
                                   REGION "GET FROM HMI"
                                       #dzLabel := #settings.viewingStation.dzData.value;
                                   END_REGION

                                   REGION "WRITE TO STATION PARAMETER"
                                       #stations.me[#i].dropZone := WSTRING_TO_USINT(#dzLabel);
                                   END_REGION

                               END_IF;
                           END_REGION

                           REGION "ON LINE LABEL INPUT"
                               IF #lineEntered THEN

                                   REGION "GET FROM HMI"
                                       #lineLabel := #settings.viewingStation.lineData.value;
                                   END_REGION

                                   REGION "WRITE TO STATION PARAMETER"
                                       #stations.me[#i].line := #lineLabel;
                                   END_REGION

                               END_IF;
                           END_REGION

                       END_IF;
                   END_REGION

               END_FOR;
           END_REGION

       END_IF;
   END_REGION
END_FUNCTION

FUNCTION "Animate Button Details" : Void   // FC19, SCL
{ S7_Optimized_Access := 'TRUE' }
VERSION : 0.1
   VAR_INPUT
      stations : "Stations";
   END_VAR
   VAR_IN_OUT
      settings : "Settings";
   END_VAR
   VAR_TEMP
      animate : USInt;
      btnCount : Int;
      btnSelected : Bool;
      deselected : USInt;
      i : Int;
      invisible : USInt;
      pBtn : Int;
      selected : USInt;
      selStnCount : Int;
      selStnNumber : Int;
   END_VAR
BEGIN
   REGION "COPY TO LOCAL"
       #btnCount := "ptsPerStn";
       #deselected := "BgGray";
       #invisible := "invisible";
       #selected := "BgLTe";
       #selStnCount := #settings.#stations.selCount;
       #selStnNumber := #settings.stations.selNumber;
   END_REGION

   REGION "ENABLE"
       IF #selStnCount >= 1 THEN

           REGION "SHOW BUTTON DETAILS"
               #animate := #deselected;
           END_REGION

       END_IF;
   END_REGION

   REGION "DISABLE"
       IF #selStnCount = 0 THEN

           REGION "HIDE BUTTON DETAILS"
               #animate := #invisible;
           END_REGION

       END_IF;
   END_REGION

   REGION "APPLY ANIMATION"
       FOR #i := 0 TO #btnCount DO

           REGION "CALCULATE BUTTON POINTER"
               #pBtn := "Pointer Calc: Button Details"(#i);
           END_REGION

           REGION "WHILE Station SELECTED"
               IF #selStnCount <> 0 THEN

                   REGION "COPY TO LOCAL"
                       #btnSelected := #stations.me[#selStnNumber].settings.btnSelection[#pBtn];
                   END_REGION

                   REGION "ANIMATE BUTTON SELECTION

                       REGION "SELECTED"
                           IF #btnSelected THEN
                               #animate := #selected;
                           END_IF;
                       END_REGION

                       REGION "NOT SELECTED"
                           IF NOT #btnSelected THEN
                               #animate := #deselected;
                           END_IF;
                       END_REGION

                   END_REGION

               END_IF;
           END_REGION


           REGION "SEND TO HMI"
               #settings.viewingStation.btns[#i].label.animate := #animate;
               #settings.viewingStation.btns[#i].alloted.animate := #animate;
               #settings.viewingStation.btns[#i].critical.animate := #animate;
               #settings.viewingStation.btns[#i].partNumber.animate := #animate;
           END_REGION

       END_FOR;
   END_REGION
END_FUNCTION

FUNCTION "Populate Station Name" : WString   // FC20, SCL
{ S7_Optimized_Access := 'TRUE' }
VERSION : 0.1
   VAR_INPUT
      line : WString;
      dropZone : USInt;
   END_VAR
BEGIN
   #"Populate Station Name" := CONCAT_WSTRING(IN1 := #line,
                                              IN2 := wstring#' ',
                                              IN3 := "Strip Sign"(USINT_TO_WSTRING(#dropZone)));
END_FUNCTION

FUNCTION "Pointer Calc: Button Details" : Int   // FC21, SCL
{ S7_Optimized_Access := 'TRUE' }
VERSION : 0.1
   VAR_INPUT
      index : Int;
   END_VAR
   VAR_TEMP
      val : Int;
   END_VAR
BEGIN
   IF #index MOD 2 = 0 THEN
       #val := 7 - #index / 2;
   END_IF;

   IF #index MOD 2 <> 0 THEN
       #val := 3 - #index / 2;
   END_IF;

   #"Pointer Calc: Button Details" := #val;
END_FUNCTION

FUNCTION "Buffer Part Req Log Row: Generate" : "Part Req Log Row"   // FC22, SCL
{ S7_Optimized_Access := 'TRUE' }
VERSION : 0.1
   VAR_INPUT
      address : Int;
      "type" : Int;
   END_VAR
   VAR_TEMP
      retVal : Int;
   END_VAR
BEGIN
   REGION "ADDRESS"
       #"Buffer Part Req Log Row: Generate".address := #address;
   END_REGION

   REGION "REQUEST TYPE"
       #"Buffer Part Req Log Row: Generate".reqType := #type;
   END_REGION

   REGION "TIME STAMP"
       #retVal := RD_SYS_T(#"Buffer Part Req Log Row: Generate".timeStamp);
   END_REGION
END_FUNCTION

FUNCTION "Sim to Global" : Void   // FC23, SCL
{ S7_Optimized_Access := 'TRUE' }
VERSION : 0.1
   VAR_INPUT
      simStations : "Simulated Stations";
   END_VAR
   VAR_IN_OUT
      stations : "Stations";
   END_VAR
   VAR_TEMP
      btnCount : Int;
      firstStn : Int;
      i : Int;
      j : Int;
      pSim : Int;
      pStn : Int;
      simKP8Count : Int;
      stnCount : Int;
   END_VAR
BEGIN
   REGION "COPY TO LOCAL"
       #btnCount := "ptsPerStn";
       #firstStn := #simStations.firstStn;
       #simKP8Count := "simKP8Count";
       #stnCount := "stnCount";
   END_REGION

   REGION "FOR EACH STATION"
       FOR #i := 0 TO #simKP8Count DO

           REGION "CALCULATE POINTER"
               #pStn := #i + #firstStn;
               #pSim := #i;
           END_REGION

           REGION "UPPER LIMIT ROLL OVER"
               IF #pStn > #stnCount THEN
                   #pStn := #firstStn + #i - #stnCount - 1;
               END_IF;
           END_REGION

           REGION "COPY SIMULATED PRESSES"
               #stations.me[#pStn].kp8In := #simStations.me[#pSim].btn.actuate;
           END_REGION

       END_FOR;
   END_REGION
END_FUNCTION

FUNCTION "Pointer Calc: KP8 Labels" : Int   // FC25, SCL
{ S7_Optimized_Access := 'TRUE' }
VERSION : 0.1
   VAR_INPUT
      index : Int;
   END_VAR
   VAR_TEMP
      val : Int;
   END_VAR
BEGIN
   IF #index >= 4 THEN
       #val := 7 - (#index - 4) * 2;
   END_IF;

   IF #index <= 3 THEN
       #val := 8 - #index * 2;
   END_IF;

   #"Pointer Calc: KP8 Labels" := #val;
END_FUNCTION

FUNCTION "KP8 Color to Sim Animation" : USInt   // FC26, SCL
{ S7_Optimized_Access := 'TRUE' }
VERSION : 0.1
   VAR_INPUT
      kp8Color : DWord;
      btnNumber : Int;
   END_VAR
   VAR_TEMP
      animate : USInt;
      blue : USInt;
      colorDWord : DWord;
      colorInt : DInt;
      green : USInt;
      off : USInt;
      red : USInt;
      white : USInt;
      yellow : USInt;
   END_VAR
   VAR CONSTANT
      blueMask : DInt := 16#0000_0100;
      btnMask : DInt := 16#0101_0100;
      greenMask : DInt := 16#0001_0000;
      offMask : DInt := 16#0000_0000;
      redMask : DInt := 16#0100_0000;
      whiteMask : DInt := 16#0101_0100;
      yellowMask : DInt := 16#0101_0000;
   END_VAR
BEGIN
   REGION "COPY TO LOCAL"
       #blue := "BgLBl";
       #green := "BgLGr";
       #off := "BgGray";
       #red := "BgLRd";
       #white := "BgWh";
       #yellow := "BgLYe";
   END_REGION

   REGION "ISOLATE BUTTON COLOR"
       #colorDWord := SHR_DWORD(IN := #kp8Color,N := INT_TO_ULINT(#btnNumber));
       #colorDWord := #colorDWord AND #btnMask;
       #colorInt := DWORD_TO_DINT(#colorDWord);
   END_REGION

   REGION "DETERMINE ANIMATION"
       CASE #colorInt OF
           #blueMask:
               #animate := #blue;
           #greenMask:
               #animate := #green;
           #redMask:
               #animate := #red;
           #whiteMask:
               #animate := #white;
           #yellowMask:
               #animate := #yellow;
           ELSE
               #animate := #off;
       END_CASE;
   END_REGION

   REGION "RETURN VALUE"
       #"KP8 Color to Sim Animation" := #animate;
   END_REGION
END_FUNCTION

FUNCTION "Recipe Nav Button" : Void   // FC32, SCL
{ S7_Optimized_Access := 'TRUE' }
VERSION : 0.1
   VAR_INPUT
      visRows : Int;
      actuate : Bool;
      maxRows : Int;
      btnNum : Int;
   END_VAR
   VAR_IN_OUT
      recipeSelectScreen : "HSS: Menu Selection Screen";
   END_VAR
   VAR_TEMP
      eval : "HSS: Menu Selection Screen";
      color : Int;
   END_VAR
BEGIN
   REGION "COPY TO LOCAL"
       #eval := #recipeSelectScreen;
   END_REGION


   REGION "NARROW"
       IF #maxRows > #visRows THEN
           #color := "BgGray";
       END_IF;
   END_REGION


   REGION "WIDE"
       IF #maxRows <= #visRows THEN
           #color := "invisible";
       END_IF;
   END_REGION


   REGION "ROW COUNT INDEPENDENT"
       IF #actuate THEN
           #color := "BgLTe";
       END_IF;
   END_REGION


   REGION "DRAW"
       #eval.animate[#btnNum] := #color;
   END_REGION


   REGION "COPY TO GLOBAL"
       #recipeSelectScreen := #eval;
   END_REGION
END_FUNCTION

FUNCTION "LRUD KP8 Remap" : Int   // FC35, SCL
{ S7_Optimized_Access := 'TRUE' }
VERSION : 0.1
   VAR_INPUT
      btnNum : Int;
      mode : Int;   // 1 = KP8; 2 = KTP700
   END_VAR
   VAR_TEMP
      output : Int;
   END_VAR
   VAR CONSTANT
      kp8 : Int := 1;
      ktp700 : Int := 2;
   END_VAR
BEGIN
   IF #btnNum >= 4 THEN
       #output := (7 - #btnNum) * 2;
   END_IF;

   IF #btnNum <= 3 THEN
       #output := (3 - #btnNum) * 2 + 1;
   END_IF;

   #"LRUD KP8 Remap" := #output;
END_FUNCTION

// folder: Unsorted/Main HMI/Network Diagnostics

FUNCTION_BLOCK "NetDiag: Get IPs"   // FB27, SCL
{ S7_Optimized_Access := 'TRUE' }
VERSION : 0.1
   VAR_OUTPUT
      error : Bool := FALSE;   // Rising edge informs that an error occurred during the execution of the FB
      status : Word := 16#0000;   // Current status of FB
      statusID : Word := 16#0;   // Current status ID of calling instruction
   END_VAR
   VAR_IN_OUT
      ioSystemData : "UserDiag_typeIOSystem";   // IO-System diagnostics data
   END_VAR
   VAR
      statError : Bool := FALSE;   // Static value for output error
      statStatus : Word := 16#0000;   // Static value for output status
      statStatusID : Word := 16#0;   // Static value for output statusID
      instGetStationInfo : GetStationInfo;   // Instance of GetStationInfo
      statFirstDeviceFlag : Bool := TRUE;   // Help tag for the first device in the linked list
      statDeviceIndex : Int := 0;   // Device/slave index
   END_VAR
   VAR_TEMP
      tempIP : IF_CONF_v4;   // Temporary IP address
   END_VAR
   VAR CONSTANT
      STATUS_EXECUTION_FINISHED : Word := 16#0000;   // Execution finished without errors
      ID_GET_STATION_INFO : Word := 12;   // StatusID during GetStationInfo command
      MODE_IPV4 : UInt := 1;   // Address parameter according to IPv4
      LAST_DEVICE : Int := -1;   // No next device
   END_VAR
BEGIN
   //=============================================================================
   //SIEMENS AG
   //(c)Copyright 2015 All Rights Reserved
   //-----------------------------------------------------------------------------
   //Library: 
   //Tested with: S7-1516-3 PN/DP FW 2.5
   //Engineering: TIA Portal V15
   //Restrictions: Call in cyclic OB
   //Requirements: -
   //Functionality: Get IP address of IO devices
   //-----------------------------------------------------------------------------
   //Change log table:
   //Version  Date       Expert in charge                Changes applied
   //01.00.00 20.12.2017 Siemens Industry Online Support First released version
   //=============================================================================

   //=============================================================================
   // Go through existing devices and get IP address
   //=============================================================================
   // Initialize the pointer for the first run 
   IF (#statFirstDeviceFlag = TRUE)
   THEN
       #statDeviceIndex := #ioSystemData.firstDevice;
       #statFirstDeviceFlag := FALSE;
   END_IF;

   // Check and store the IP address, if the device is existing
   // GetStationInfo is an acyclic instruction. In the FB, the
   // instruction has to be repeated until it is done or error
   IF ((#ioSystemData.number >= 100)
       AND (#ioSystemData.number <= 115)
       AND (#ioSystemData.devices[#statDeviceIndex].exists = TRUE)
       AND (#ioSystemData.devices[#statDeviceIndex].ipAddress.ADDR[1] = 0))
   THEN
       // Get IP address of each decive in PN System
       #instGetStationInfo(REQ := TRUE,
                           LADDR := #ioSystemData.devices[#statDeviceIndex].hardwareId,
                           MODE := #MODE_IPV4,
                           DATA := #tempIP);

       IF (#instGetStationInfo.ERROR = TRUE)
       THEN
           // Error handling
           #statStatus := #instGetStationInfo.STATUS;
           #statStatusID := #ID_GET_STATION_INFO;
           #statError := TRUE;

           // Everything is ok --> Copy IP address    
       ELSIF (#instGetStationInfo.DONE = TRUE)
       THEN
           #ioSystemData.devices[#statDeviceIndex].ipAddress := #tempIP.InterfaceAddress;

           // Initialize the pointer for the next run
           #statDeviceIndex := #ioSystemData.devices[#statDeviceIndex].nextDevice;
       ELSE
           ;
       END_IF;
   ELSE
       // Initialize the pointer for the next run
       #statDeviceIndex := #ioSystemData.devices[#statDeviceIndex].nextDevice;
   END_IF;

   // Check last device
   IF (#statDeviceIndex = #LAST_DEVICE)
   THEN
       #statDeviceIndex := #ioSystemData.firstDevice;
   END_IF;

   // Write static values to outputs
   #error := #statError;
   #status := #statStatus;
   #statusID := #statStatusID;
END_FUNCTION_BLOCK

FUNCTION_BLOCK "NetDiag: Coordinate"   // FB28, LAD
{ S7_Optimized_Access := 'TRUE' }
VERSION : 0.1
// //============================================================================
// //SIEMENS AG
// //(c)Copyright 2017 All Rights Reserved
// //-----------------------------------------------------------------------------
// //Library: -
// //Tested with: S7-1516-3 PN/DP FW 2.5
// //Engineering: TIA Portal V15
// //Restrictions: -
// //Requirements: -
// //Functionality: Main FB for diagnostics
// //-----------------------------------------------------------------------------
// //Change log table:
// //Version  Date              Expert in charge                               Changes applied
// //01.00.00 25.04.2017 Siemens Industry Online Support First released version
// //01.01.00 01.12.2017 Siemens Industry Online Support Renamed in "UserDiag_Diagnostics"
// //                                                                                                    Check Flag "startDiag"
// //============================================================================
   VAR_IN_OUT
      startDiag : Bool := false;   // Startflag for diagnostic
      plcData : "UserDiag_typePLC";   // PLC diagnostics data
      ioSystemData : Array[1.."USERDIAG_IO_SYSTEMS_UPPER_LIM"] of "UserDiag_typeIOSystem";   // IO-System diagnostics data
   END_VAR
   VAR
      instPLCChk : "NetDiag: Check PLC";   // Instance of "UserDiag_PLCCheck"
      instIOSysChk : "NetDiag: IO Systems";   // Instance of "UserDiag_IOSystemCheck"
   END_VAR
BEGIN

REGION Network 1: Check Startflag for diagnostic
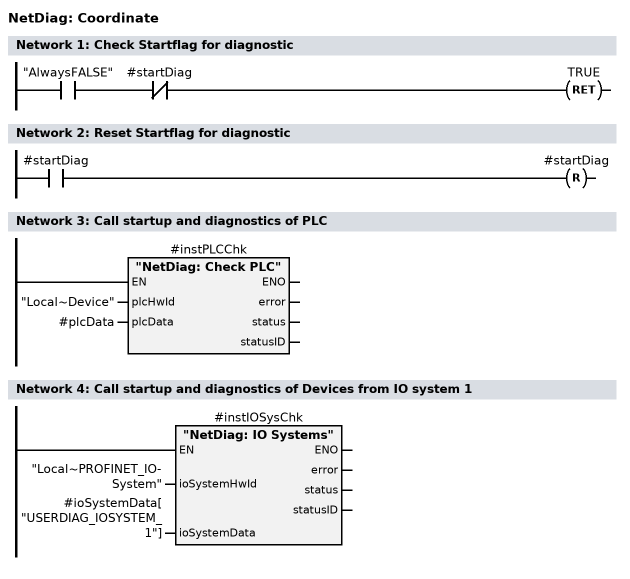
   IF "AlwaysFALSE" AND NOT #startDiag THEN
       ENO := TRUE;
       RETURN;
   END_IF;
END_REGION

REGION Network 2: Reset Startflag for diagnostic
   RUNG wire#powerrail
      Contact( #startDiag )
      R_Coil( #startDiag )
   END_RUNG
   // the same network as SCL:
   IF #startDiag THEN #startDiag := FALSE; END_IF;
END_REGION

REGION Network 3: Call startup and diagnostics of PLC
   RUNG wire#powerrail
      #instPLCChk(plcHwId := "Local~Device", plcData := #plcData, error =>, status =>, statusID =>)
   END_RUNG
   // the same network as SCL:
   #instPLCChk(plcHwId := "Local~Device", plcData := #plcData);   // "NetDiag: Check PLC"
END_REGION

REGION Network 4: Call startup and diagnostics of Devices from IO system 1
   RUNG wire#powerrail
      #instIOSysChk(ioSystemHwId := "Local~PROFINET_IO-System", ioSystemData := #ioSystemData["USERDIAG_IOSYSTEM_1"], error =>, status =>, statusID =>)
   END_RUNG
   // the same network as SCL:
   #instIOSysChk(ioSystemHwId := "Local~PROFINET_IO-System",   // "NetDiag: IO Systems"
                 ioSystemData := #ioSystemData["USERDIAG_IOSYSTEM_1"]);
END_REGION
END_FUNCTION_BLOCK

FUNCTION_BLOCK "NetDiag: Check PLC"   // FB29, SCL
{ S7_Optimized_Access := 'TRUE' }
VERSION : 0.1
   VAR_INPUT
      plcHwId : Hw_Device := 0;   // Hardware ID
   END_VAR
   VAR_OUTPUT
      error : Bool := FALSE;   // Rising edge informs that an error occurred during the execution of the FB
      status : Word := 16#0000;   // Current status of FB
      statusID : Word := 16#0;   // Current status ID of calling instruction
   END_VAR
   VAR_IN_OUT
      plcData : "UserDiag_typePLC";   // PLC diagnostics data
   END_VAR
   VAR
      statError : Bool := FALSE;   // Static value for output error
      statStatus : Word := 16#0000;   // Static value for output status
      statStatusID : Word := 16#0;   // Static value for output statusID
      statGeoAddr : GEOADDR;   // Slot information
      statGeoLaddr : Hw_Any := 16#0000;   // GEO2LOG hardware identifier
      statProblemPlcModulStates : Array[0..#MODULES_STATES_UPPER_LIM] of Bool;   // Storage of the status of all modules in the PLC central station --> State: Problem
      statFaultyPlcModulStates : Array[0..#MODULES_STATES_UPPER_LIM] of Bool;   // Storage of the status of all modules in the PLC central station --> State: Faulty
      statExistingPlcModulStates : Array[0..#MODULES_STATES_UPPER_LIM] of Bool;   // Storage of the status of all modules in the PLC central station --> State: Exists
      statActualCentralModules : USInt := 0;   // Actual number of modules in the central station (PLC)
   END_VAR
   VAR_TEMP
      tempSlotNum : Int;   // Index slot number
      tempRetValGeo : Int;   // GEO2LOG error information
      tempRetValModuleStates : Int;   // Return value system function ModuleStates
   END_VAR
   VAR CONSTANT
      STATUS_EXECUTION_FINISHED : Word := 16#0000;   // Execution finished without errors
      ERR_MAX_SLOTS_PER_PLC : Word := 16#8400;   // There are more modules configured as defined with the user constant: USERDIAG_SLOTS_PER_PLC_UPPER_LIM
      ID_LOCAL : Word := 1;   // StatusID local
      ID_MODULE_STATES_CONFIGURED : Word := 2;   // StatusID during ModuleStates command (configured mode)
      ID_MODULE_STATES_FAULTY : Word := 3;   // StatusID during ModuleStates command (faulty mode)
      ID_MODULE_STATES_PROBLEM : Word := 4;   // StatusID during ModuleStates command (problem mode)
      ID_MODULE_STATES_EXISTING : Word := 5;   // StatusID during ModuleStates command (existing mode)
      ID_LED : Word := 12;   // StatusID occurred during LED command
      MODE_FAULTY : USInt := 2;   // Used for instruction DeviceStates, read out all faulty devices
      MODE_EXIST : USInt := 4;   // Used for instruction DeviceStates, read out all devices not reachable
      MODE_PROBLEM : USInt := 5;   // Used for instruction DeviceStates, read out all devices with several problems
      STATE_OK : USInt := 1;   // Module state: ok
      STATE_FAULT : USInt := 2;   // Modulestate: fault
      STATE_PROBLEM : USInt := 5;   // Module state: problem
      STATE_WAS_FAULT : USInt := 12;   // Module state: was fault
      STATE_PROBLEM_GONE : USInt := 15;   // Module state: had a problem
      MODULE_OF_PLC : USInt := 4;   // GEO2LOG structure: HW type = 4
      CPU : USInt := 0;   // GEO2LOG structure: Area = 0
      CENTRAL_SYSTEM : USInt := 0;   // GEO2LOG structure: IO System = 0
      CENTRAL_STATION : USInt := 0;   // GEO2LOG structure: Station = 0
      NO_LED : Int := 0;   // LED does not exist
      LED_OFF : Int := 1;   // LED is permanently switched off
      LED_NO_INFO : Int := 9;   // LED exists, but status information not available
      MODULES_STATES_UPPER_LIM : Int := 127;   // Upper array limit for output tag of instruction ModuleStates
      ERROR_LED : UInt := 2;   // Identification number of the LED
   END_VAR
BEGIN
   //=============================================================================
   //SIEMENS AG
   //(c)Copyright 2017 All Rights Reserved
   //-----------------------------------------------------------------------------
   //Library: 
   //Tested with: S7-1516-3 PN/DP FW 2.5
   //Engineering: TIA Portal V15
   //Restrictions: Call in cyclic OB
   //Requirements: -
   //Functionality: Determine plc state and local module states
   //-----------------------------------------------------------------------------
   //Change log table:
   //Version  Date       Expert in charge                Changes applied
   //01.00.00 27.01.2017 Siemens Industry Online Support First released version
   //01.00.01 20.12.2017 Siemens Industry Online Support actualConfiguredSlots >= 1
   //01.00.02 27.02.2018 Siemens Industry Online Support Minor corrections
   //=============================================================================

   IF (#plcData.hardwareId = 0)
   THEN
       #statGeoAddr.HWTYPE := #MODULE_OF_PLC;      // Hardware type 4: module
       #statGeoAddr.AREA := #CPU;                  // Area ID 0: CPU
       #statGeoAddr.IOSYSTEM := #CENTRAL_SYSTEM;   // PROFINET IO system (0 = central unit in the rack)
       #statGeoAddr.STATION := #CENTRAL_STATION;   // Number of the rack if area identifier AREA = 0 (central module)

       #statStatus := #STATUS_EXECUTION_FINISHED;
       #statStatusID := 0;
       #statError := FALSE;
       #statActualCentralModules := 0;

       FOR #tempSlotNum := 0 TO "USERDIAG_SLOTS_PER_PLC_UPPER_LIM" DO
           // Slot number
           #statGeoAddr.SLOT := INT_TO_UINT(#tempSlotNum);
           // read LADDR from local modules
           #tempRetValGeo := GEO2LOG(GEOADDR := #statGeoAddr,
                                     LADDR => #statGeoLaddr);
           // Check Retval
           IF ((#tempRetValGeo = 0)
               AND (#statGeoLaddr <> 16#0))
           THEN
               // Store LADDR from local modules in diagnostic data block
               IF (#tempSlotNum = 1)
               THEN
                   #plcData.hardwareId := #statGeoLaddr;
               END_IF;
               #plcData.slots[#tempSlotNum].hardwareId := #statGeoLaddr;
               #statActualCentralModules := #statActualCentralModules + 1;
               #plcData.slots[#tempSlotNum].configured := TRUE;
           ELSE
               // If the return value ist not = 0 --> the device/system/module is not
               // configured --> No error handling
               // set LADDR from local modules to 0 in diagnostic data block
               #plcData.slots[#tempSlotNum].hardwareId := 0;
               #plcData.slots[#tempSlotNum].configured := FALSE;
           END_IF;
           // Store the actual configured devices in the diagnostics DB
           #plcData.actualConfiguredSlots := #statActualCentralModules;
       END_FOR;

       // Check if further slots are configured
       #statGeoAddr.SLOT := INT_TO_UINT(#tempSlotNum);

       #tempRetValGeo := GEO2LOG(GEOADDR := #statGeoAddr,
                                 LADDR => #statGeoLaddr);

       IF ((#tempRetValGeo = 0)
           AND (#statGeoLaddr <> 16#0))
       THEN
           // In the PLC are more slots configured as defined with the user constant
           #statStatus := #ERR_MAX_SLOTS_PER_PLC;
           #statStatusID := #ID_LOCAL;
           #statError := TRUE;
       END_IF;

   END_IF;

   // Reset PLC error state
   #plcData.error := FALSE;

   //=============================================================================
   // Check modul states from LOCAL MODULES
   //=============================================================================
   // Check if central module are available - at least one module is always
   // configured, the PLC itself
   IF (#plcData.actualConfiguredSlots >= 1)
   THEN

       // Check the status of the local modules
       #tempRetValModuleStates := ModuleStates(LADDR := #plcHwId,
                                               MODE := #MODE_PROBLEM,
                                               STATE := #statProblemPlcModulStates);

       // Check if the block call was successful
       IF (#tempRetValModuleStates <> 0)
       THEN
           // Error handling
           #statStatus := INT_TO_WORD(#tempRetValModuleStates);
           #statStatusID := #ID_MODULE_STATES_PROBLEM;
           #statError := TRUE;
       ELSE
           ; // Everything is ok!
       END_IF;

       #tempRetValModuleStates := ModuleStates(LADDR := #plcHwId,
                                               MODE := #MODE_FAULTY,
                                               STATE := #statFaultyPlcModulStates);

       // Check if the block call was successful
       IF (#tempRetValModuleStates <> 0)
       THEN
           // Error handling
           #statStatus := INT_TO_WORD(#tempRetValModuleStates);
           #statStatusID := #ID_MODULE_STATES_FAULTY;
           #statError := TRUE;
       ELSE
           ; // Everything is ok!
       END_IF;

       #tempRetValModuleStates := ModuleStates(LADDR := #plcHwId,
                                               MODE := #MODE_EXIST,
                                               STATE := #statExistingPlcModulStates);

       // Check if the block call was successful
       IF (#tempRetValModuleStates <> 0)
       THEN
           // Error handling
           #statStatus := INT_TO_WORD(#tempRetValModuleStates);
           #statStatusID := #ID_MODULE_STATES_EXISTING;
           #statError := TRUE;
       ELSE
           ; // Everything is ok!
       END_IF;

   ELSE
       ; // There are no central moduls configured
   END_IF;

   //=============================================================================
   // Set module states of LOCAL MODULES
   //=============================================================================
   #tempSlotNum := 0;
   WHILE (#tempSlotNum <= #plcData.actualConfiguredSlots)
   DO
       IF (#plcData.slots[#tempSlotNum].configured)
       THEN
           IF (#statExistingPlcModulStates[#tempSlotNum + 1] = TRUE)
           THEN
               #plcData.slots[#tempSlotNum].exists := TRUE;
               CASE #plcData.slots[#tempSlotNum].state OF
                   #STATE_WAS_FAULT,
                   #STATE_PROBLEM_GONE:
                       ;
                   #STATE_FAULT:
                       #plcData.slots[#tempSlotNum].state := #STATE_WAS_FAULT;
                   #STATE_PROBLEM:
                       #plcData.slots[#tempSlotNum].state := #STATE_PROBLEM_GONE;
                   ELSE
                       #plcData.slots[#tempSlotNum].state := #STATE_OK;
               END_CASE;
           ELSE
               #plcData.slots[#tempSlotNum].error := TRUE;
               #plcData.error := TRUE;
               #plcData.slots[#tempSlotNum].exists := FALSE;
           END_IF;

           IF (#statFaultyPlcModulStates[#tempSlotNum + 1] = TRUE)
           THEN
               // Modul is faulty
               #plcData.slots[#tempSlotNum].faulty := TRUE;
               #plcData.slots[#tempSlotNum].problem := TRUE;
               #plcData.slots[#tempSlotNum].error := TRUE;
               #plcData.slots[#tempSlotNum].state := #STATE_FAULT;
           ELSIF (#statProblemPlcModulStates[#tempSlotNum + 1] = TRUE)
           THEN
               // Modul has a problem
               #plcData.slots[#tempSlotNum].faulty := FALSE;
               #plcData.slots[#tempSlotNum].problem := TRUE;
               #plcData.slots[#tempSlotNum].error := TRUE;
               #plcData.slots[#tempSlotNum].state := #STATE_PROBLEM;
           ELSE
               // Modul is OK
               #plcData.slots[#tempSlotNum].error := FALSE;
               #plcData.slots[#tempSlotNum].problem := FALSE;
               #plcData.slots[#tempSlotNum].faulty := FALSE;
           END_IF;

           // Error in PLC - Slot = 1, but index must be increased by 1, because of bit 0 = group display
           // --> used index = 2
           IF (#statProblemPlcModulStates[2] = TRUE)
               OR (#statFaultyPlcModulStates[2] = TRUE)
           THEN
               #plcData.error := TRUE;
           END_IF;
       END_IF;

       #tempSlotNum := #tempSlotNum + 1;
   END_WHILE;

   // Write static values to outputs
   #error := #statError;
   #status := #statStatus;
   #statusID := #statStatusID;

   //----------------------------------------------------------------------------------------------
END_FUNCTION_BLOCK

FUNCTION_BLOCK "NetDiag: IO Systems"   // FB30, SCL
{ S7_Optimized_Access := 'TRUE' }
VERSION : 0.1
   VAR_INPUT
      ioSystemHwId : Hw_IoSystem := 16#0000;   // This ID is representing the IO System (PN or DP), find the ID in the system constants
   END_VAR
   VAR_OUTPUT
      error : Bool := FALSE;   // Rising edge informs that an error occurred during the execution of the FB
      status : Word := 16#0000;   // Current status of FB
      statusID : Word := 16#0;   // Current status ID of calling instruction
   END_VAR
   VAR_IN_OUT
      ioSystemData : "UserDiag_typeIOSystem";   // IO-System diagnostics data
   END_VAR
   VAR
      statError : Bool := FALSE;   // Static value for output error
      statStatus : Word := 16#0000;   // Static value for output status
      statStatusID : Word := 16#0;   // Static value for output statusID
      statActualConfiguredDevices : Int := 0;   // Actual number of devices/slaves in the IOSystem/DP-Mastersystem
      statGeoAddr : GEOADDR;   // Slot information
      statGeoLaddr : Hw_Any := 16#0000;   // GEO2LOG hardware identifier
      statConfiguredDevices : Array[0..#DEVICES_STATES_UPPER_LIM] of Bool;   // Temporary storage of the return of "DeviceStates", to combine the states of the devices/slaves with numbers and names
      statExistingDevices : Array[0..#DEVICES_STATES_UPPER_LIM] of Bool;   // Temporary storage of the return of "DeviceStates", to combine the states of the devices/slaves with numbers and names
      statFaultyDevices : Array[0..#DEVICES_STATES_UPPER_LIM] of Bool;   // Temporary storage of the return of "DeviceStates", to combine the states of the devices/slaves with numbers and names
      statDisabledDevices : Array[0..#DEVICES_STATES_UPPER_LIM] of Bool;   // Temporary storage of the return of "DeviceStates", to combine the states of the devices/slaves with numbers and names
      statProblemDevices : Array[0..#DEVICES_STATES_UPPER_LIM] of Bool;   // Temporary storage of the return of "DeviceStates", to combine the states of the devices/slaves with numbers and names
      statDeviceProblemModules : Array[0..#MODULES_STATES_UPPER_LIM] of Bool;   // Storage of the status of all modules in the PN Devices / PB Slaves --> State: Problem
      statDeviceFaultyModules : Array[0..#MODULES_STATES_UPPER_LIM] of Bool;   // Storage of the status of all modules in the PN Devices / PB Slaves --> State: Faulty
      statDeviceExistingModules : Array[0..#MODULES_STATES_UPPER_LIM] of Bool;   // Storage of the status of all modules in the PN Devices / PB Slaves --> State: Existing
      instGetNameDevices : Get_Name;   // Instance of the system function "GetName"
      statInitString : String := '';   // Used to initialize the temporary string to convert into STRING[50]
      statFirstDevice : UInt := 0;   // Station number of the first device of the list
      statFirstDeviceFlag : Bool := TRUE;   // Help tag for the first device in the linked list
      statLastDevice : UInt := 0;   // Station number of the last device of the list
      statMaxDevices : Int := 0;   // Max devices per IO system
   END_VAR
   VAR_TEMP
      tempIndex : Int;   // Index of configured devices/slaves
      tempDeviceIndex : Int;   // Device/slave index
      tempSlotIndex : Int;   // Slot index
      tempSlotNum : Int;   // Index module number
      tempRetValGeo : Int;   // GEO2LOG error information
      tempRetValDeviceStates : Int;   // DeviceStates error information
      tempRetValModuleStates : Int;   // Return value of the system function "ModuleStates"
      tempStringConvert : String;   // Store the device names temporary here, to convert them into STRING[50]
      tempLastDevice : UInt;   // Temporary storage of the actual index, if it´s the last device --> store it in static
      tempDeviceInit : "UserDiag_typeDevice";   // Initalization of the device/slave diagnostic structure
   END_VAR
   VAR CONSTANT
      STATUS_EXECUTION_FINISHED : Word := 16#0000;   // Execution finished without errors
      ERR_MAX_SLOTS_PER_DEVICE : Word := 16#8400;   // There are more modules configured as defined with the user constant: USERDIAG_SLOTS_PER_DEVICE_UPPER_LIM
      ERR_MAX_DEVICES_PER_IOSYSTEM : Word := 16#8401;   // There are more modules configured as defined with the user constant: USERDIAG_DEVICES_PER_IO_SYTEM_UPPER_LIM
      ID_LOCAL : Word := 1;   // StatusID local
      ID_MODULE_STATES_CONFIGURED : Word := 2;   // StatusID during ModuleStates command (configured mode)
      ID_MODULE_STATES_FAULTY : Word := 3;   // StatusID during ModuleStates command (faulty mode)
      ID_MODULE_STATES_PROBLEM : Word := 4;   // StatusID during ModuleStates command (problem mode)
      ID_MODULE_STATES_EXISTING : Word := 5;   // StatusID during ModuleStates command (existing mode)
      ID_DEVICE_STATES_CONFIGURED : Word := 6;   // StatusID during DeviceStates command (configuration mode)
      ID_DEVICE_STATES_FAULTY : Word := 7;   // StatusID during DeviceStates command (fault mode)
      ID_DEVICE_STATES_PROBLEM : Word := 8;   // StatusID during DeviceStates command (problem mode)
      ID_DEVICE_STATES_EXISTING : Word := 9;   // StatusID during DeviceStates command (existing mode)
      ID_DEVICE_STATES_DISABLED : Word := 10;   // StatusID during DeviceStates command (disable mode)
      ID_GET_NAME : Word := 11;   // StatusID during GET_NAME command
      MODE_CONFIGURED : USInt := 1;   // Used for instruction DeviceStates/ModuleStates, read out all configured devices/slaves
      MODE_FAULTY : USInt := 2;   // Used for instruction DeviceStates/ModuleStates, read out all faulty devices/slaves
      MODE_DISABLED : USInt := 3;   // Used for instruction DeviceStates/ModuleStates, read out all disabled devices/slaves
      MODE_EXIST : USInt := 4;   // Used for instruction DeviceStates/ModuleStates, read out all devices/slaves not reachable
      MODE_PROBLEM : USInt := 5;   // Used for instruction DeviceStates/ModuleStates, read out all devices with several problems
      DEVICE_SLAVE : USInt := 2;   // GEO2LOG structure: HW type = 2
      MODULE_OF_DEVICE : USInt := 4;   // GEO2LOG structure: HW type = 4
      IO_SYSTEM_AREA : USInt := 1;   // GEO2LOG structure: Area = 1
      DP_SYSTEM_AREA : USInt := 2;   // GEO2LOG structure: Area = 2
      STATE_OK : USInt := 1;   // Device/modul state: ok
      STATE_FAULT : USInt := 2;   // Device/modul state: fault
      STATE_LOST_CON : USInt := 3;   // Device/modul state: lost connection
      STATE_DISABLED : USInt := 4;   // Device/modul state: disabled
      STATE_PROBLEM : USInt := 5;   // Device/modul state: problem
      STATE_WAS_FAULT : USInt := 12;   // Device/modul state: was fault
      STATE_WAS_LOST : USInt := 13;   // Device/modul state: connection was lost
      STATE_WAS_DISABLED : USInt := 14;   // Device/modul state: device/slave was disabled
      STATE_PROBLEM_GONE : USInt := 15;   // Device/modul state: had a problem
      MODULES_STATES_UPPER_LIM : Int := 127;   // Upper array limit for output tag of instruction ModuleStates
      DEVICES_STATES_UPPER_LIM : Int := 1023;   // Upper array limit for output tag of instruction DeviceStates
      ERR_HWID_NOT_EXISTENT : Int := 16#8091;   // Hardware identifier of the LADDR parameter does not exist. Check (for example, in the system constants) whether the value for LADDR exists in the project.
      ERR_LADDR_ADDRESS : Int := 16#8092;   // LADDR does not address a PROFINET IO or DP master system.
      POS_FIRST_CHAR : Int := 50;   // Position of first character to be deleted
      NUMBER_CHAR : Int := 204;   // Number of characters to be deleted
      MAX_SLAVES_DP : Int := 127;   // Max number of slaves in a PROFIBUS IO system
      LAST_DEVICE : Int := -1;   // No next device
   END_VAR
BEGIN
   //=============================================================================
   //SIEMENS AG
   //(c)Copyright 2015 All Rights Reserved
   //-----------------------------------------------------------------------------
   //Library: 
   //Tested with: S7-1516-3 PN/DP FW 2.5
   //Engineering: TIA Portal V15
   //Restrictions: Call in cyclic OB
   //Requirements: -
   //Functionality: Determine hardware identifier and module states from local and
   //               device modules 
   //-----------------------------------------------------------------------------
   //Change log table:
   //Version  Date       Expert in charge                Changes applied
   //01.00.00 27.01.2017 Siemens Industry Online Support First released version
   //01.00.01 20.12.2017 Siemens Industry Online Support GetStationInfo removed
   //01.00.02 27.02.2018 Siemens Industry Online Support Minor corrections
   //=============================================================================

   IF (#ioSystemHwId <> #ioSystemData.hardwareId)
   THEN
       // New IO System detected at input
       #statFirstDeviceFlag := TRUE;
       #statFirstDevice := 1;
       #statLastDevice := 1;

       #statActualConfiguredDevices := 0;
       #tempDeviceIndex := 1;

       #statError := FALSE;
       #statStatus := #STATUS_EXECUTION_FINISHED;
       #statStatusID := 0;
       #ioSystemData.error := FALSE;
       #ioSystemData.hardwareId := #ioSystemHwId;

       // Find out the number of the assigned IO system
       #tempRetValGeo := LOG2GEO(LADDR := #ioSystemHwId,
                                 GEOADDR := #statGeoAddr);
       // Set IO system ID
       #ioSystemData.number := #statGeoAddr.IOSYSTEM;

       // Initialize the structure for system function GEO2LOG
       #statGeoAddr.HWTYPE := #DEVICE_SLAVE;   // Hardware type 2: IO device

       // Predefine the type OF IO system. Either Profinet IO or Profibus DP
       IF (#statGeoAddr.AREA = #IO_SYSTEM_AREA)     // Area ID 1: PROFINET IO
       THEN
           #statMaxDevices := "USERDIAG_DEVICES_PER_IO_SYSTEM_UPPER_LIM";
       ELSIF (#statGeoAddr.AREA = #DP_SYSTEM_AREA) // Area ID 2: Profibus DP
       THEN
           IF ("USERDIAG_DEVICES_PER_IO_SYSTEM_UPPER_LIM" > #MAX_SLAVES_DP)
           THEN
               #statMaxDevices := #MAX_SLAVES_DP;
           ELSE
               #statMaxDevices := "USERDIAG_DEVICES_PER_IO_SYSTEM_UPPER_LIM";
           END_IF;
       ELSE
           #statMaxDevices := "USERDIAG_DEVICES_PER_IO_SYSTEM_UPPER_LIM";
       END_IF;

       // Set all other devices to not configured
       FOR #tempIndex := 1 TO "USERDIAG_DEVICES_PER_IO_SYSTEM_UPPER_LIM" DO
           #ioSystemData.devices[#tempIndex] := #tempDeviceInit;
       END_FOR;

       //=============================================================================
       // CONFIGURED DEVICES
       //=============================================================================
       // Find out how much devices are configured in the IO System --> PROFINET IO
       // This number is the maximum number of devices, which will be checked in the
       // following programm
       #tempRetValDeviceStates := DeviceStates(LADDR := #ioSystemHwId,
                                               MODE := #MODE_CONFIGURED,
                                               STATE := #statConfiguredDevices);

       // Check if the block call was successful
       IF (#tempRetValDeviceStates = 0)
       THEN
           // Call ok
           ;
       ELSIF (#tempRetValDeviceStates = #ERR_HWID_NOT_EXISTENT)
           OR (#tempRetValDeviceStates = #ERR_LADDR_ADDRESS)
       THEN
           #ioSystemData.error := TRUE;
           #statStatus := INT_TO_WORD(#tempRetValDeviceStates);
           #statStatusID := #ID_DEVICE_STATES_CONFIGURED;
           #statError := TRUE;
       ELSE
           // Error handling
           #statStatus := INT_TO_WORD(#tempRetValDeviceStates);
           #statStatusID := #ID_DEVICE_STATES_CONFIGURED;
           #statError := TRUE;
       END_IF;

       // Check if further devices are configured
       FOR #tempIndex := 1 TO #DEVICES_STATES_UPPER_LIM DO
           IF (((#statConfiguredDevices[#tempIndex] = TRUE)
               AND (#tempIndex > #statMaxDevices))
               AND (
               ((#statGeoAddr.AREA = #DP_SYSTEM_AREA)
               AND (#tempIndex < #MAX_SLAVES_DP))
               OR (#statGeoAddr.AREA = #IO_SYSTEM_AREA))
               )
           THEN
               // In the IOSystem are more devices configured as defined with the user constant
               #statStatus := #ERR_MAX_DEVICES_PER_IOSYSTEM;
               #statStatusID := #ID_LOCAL;
               #statError := TRUE;
           END_IF;
       END_FOR;

       //=============================================================================
       // Go trough all devices and get the status of the configured
       //=============================================================================
       FOR #tempIndex := 1 TO #statMaxDevices DO
           // The devices are configured --> Read out the logical address and the
           // device name
           IF (#statConfiguredDevices[#tempIndex] = TRUE)
           THEN
               // Store the first configured device for the linked list
               IF (#statFirstDeviceFlag = TRUE)
               THEN
                   #statFirstDevice := INT_TO_UINT(#tempIndex);
                   #ioSystemData.firstDevice := UINT_TO_INT(#statFirstDevice);
                   #statFirstDeviceFlag := FALSE;
                   #tempLastDevice := INT_TO_UINT(#tempIndex);
                   // It´s not the first bit --> Store the actual index as "next device"
                   // in the further one!
               ELSE
                   #ioSystemData.devices[#tempLastDevice].nextDevice := #tempIndex;
                   #tempLastDevice := INT_TO_UINT(#tempIndex);
               END_IF;
               // Store the index of the last device for the exit condition of the
               // followiing instructions
               #statLastDevice := #tempLastDevice;
               #ioSystemData.lastDevice := UINT_TO_INT(#statLastDevice);

               // Initialize the structure for system function GEO2LOG
               #statGeoAddr.STATION := INT_TO_UINT(#tempIndex); // Station number 
               #statGeoAddr.HWTYPE := #DEVICE_SLAVE;   // Hardware type 2: IO device

               // Read LADDR from devices
               #tempRetValGeo := GEO2LOG(GEOADDR := #statGeoAddr,
                                         LADDR => #statGeoLaddr);
               // Everything is ok!
               IF (#tempRetValGeo = 0)
               THEN
                   // Store LADDR from devices in diagnostics data block
                   #ioSystemData.devices[#tempIndex].hardwareId := #statGeoLaddr;
                   #ioSystemData.devices[#tempIndex].number := INT_TO_UINT(#tempIndex);
                   #ioSystemData.devices[#tempIndex].configured := TRUE;

                   // Store the device name, if the device is existing
                   // Get name is an acyclic instruction. In the startup OB, the
                   // instruction has to be repeated until it is done or error
                   REPEAT
                       // Get device name of each decive in PN System
                       #instGetNameDevices(LADDR := #ioSystemHwId,
                                           STATION_NR := #statGeoAddr.STATION,
                                           DATA := #tempStringConvert);

                   UNTIL ((#instGetNameDevices.DONE = TRUE)
                       OR (#instGetNameDevices.ERROR = TRUE))
                   END_REPEAT;

                   IF (#instGetNameDevices.ERROR = TRUE)
                   THEN
                       // Error handling
                       #statStatus := #instGetNameDevices.STATUS;
                       #statStatusID := #ID_GET_NAME;
                       #statError := TRUE;

                       // Everything is ok --> Convert the String[254] into String[50]    
                   ELSIF (#instGetNameDevices.DONE = TRUE)
                   THEN
                       // Cut all characters more than 50 to reduce the string length
                       #ioSystemData.devices[#tempIndex].name := STRING_TO_WSTRING(DELETE(IN := #tempStringConvert,
                                                                                          L := #NUMBER_CHAR,
                                                                                          P := #POS_FIRST_CHAR));

                       // Initialize the temporary string before next loop
                       #tempStringConvert := #statInitString;
                   ELSE
                       ;
                   END_IF;


                   //=============================================================================
                   // Get the logical address of all modules and store the actual number of
                   // modules from each device
                   //=============================================================================

                   // Initialize the structure for system function GEO2LOG
                   #statGeoAddr.HWTYPE := #MODULE_OF_DEVICE;   // Hardware type 4: Module

                   FOR #tempSlotNum := 0 TO "USERDIAG_SLOTS_PER_DEVICE_UPPER_LIM" DO
                       // Slot number
                       #statGeoAddr.SLOT := INT_TO_UINT(#tempSlotNum);
                       // read LADDR from modules
                       #tempRetValGeo := GEO2LOG(GEOADDR := #statGeoAddr,
                                                 LADDR => #statGeoLaddr);
                       // check Retval
                       IF (#tempRetValGeo = 0)
                       THEN
                           // Store LADDR from modules in diagnostic data block
                           #ioSystemData.devices[#tempIndex].slots[#tempSlotNum].hardwareId := #statGeoLaddr;
                           #ioSystemData.devices[#tempIndex].actualConfiguredSlots := #ioSystemData.devices[#tempIndex].actualConfiguredSlots + 1;

                           #ioSystemData.devices[#tempIndex].slots[#tempSlotNum].configured := TRUE;

                       ELSE
                           // If the return value is not 0 --> the device/system/module is
                           // not configured --> No error handling
                           // set LADDR from modules to 0 in diagnostic data block
                           #ioSystemData.devices[#tempIndex].slots[#tempSlotNum].hardwareId := 0;
                       END_IF;
                   END_FOR;

                   // Check if further slots are configured
                   #statGeoAddr.SLOT := INT_TO_UINT(#tempSlotNum);

                   #tempRetValGeo := GEO2LOG(GEOADDR := #statGeoAddr,
                                             LADDR => #statGeoLaddr);

                   IF ((#tempRetValGeo = 0)
                       AND (#statGeoLaddr <> 16#0))
                   THEN
                       // In the PLC are more slots configured as defined with the user constant
                       #statStatus := #ERR_MAX_SLOTS_PER_DEVICE;
                       #statStatusID := #ID_LOCAL;
                       #statError := TRUE;
                   END_IF;

                   // Increment the actual configured devices, store the state and
                   // HW_ID as an numerical value (UINT)
                   #statActualConfiguredDevices := #statActualConfiguredDevices + 1;
               ELSE
                   ;
               END_IF;

           ELSE
               ; // Device not configured
           END_IF;
       END_FOR;

       #ioSystemData.actualConfiguredDevices := #statActualConfiguredDevices;

       // Mark parameter "Next Device" of the last device in the list
       // --> "Next Device" = negative --> Last device in the list
       #ioSystemData.devices[#statLastDevice].nextDevice := #LAST_DEVICE;

   END_IF; // New IO System detected at input

   #ioSystemData.error := FALSE; // Reset the IO-System error status


   //=============================================================================
   // START DIAGNOSTICS EVALUATION
   //=============================================================================

